// Mitsubishi GX Works2 project: ZhaoQing_OCV__Debug   PLC: Q10UDEH (continued)

Conveyor12109(ConveyorMotor:=ConveyorIO12109);
ConveyorIO12109.xForward:=M53;
ConveyorIO12109.xCWPresent:=X29;
Y22A:=ConveyorIO12109.xMotorCW;
M326:=NOT ConveyorIO12109.xEmpty;
M327:=ConveyorIO12109.xError;
ConveyorIO12109.iDeviceID:=12109;

Switch12310(ConveyorEntryIO:=ConveyorIO12110 ,
                                                        ConveyorExitIO:=ConveyorIO12117 ,
                                                        SwitchIO:=SwitchIO12310 );
SwitchIO12310.xLiftCylinderExtendButton:=M54;
SwitchIO12310.xLiftCylinderRetractButton:=M55;
Y22E:=SwitchIO12310.xLiftCylinderExtend;
Y22D:=SwitchIO12310.xLiftCylinderRetract;
SwitchIO12310.xLiftCylinderExtendDetect:=X2D;
SwitchIO12310.xLiftCylinderRetractDetect:=X2E;
ConveyorIO12110.xForward:=M56;
ConveyorIO12110.xCWPresent:=X2F OR X30;
Y22C:=ConveyorIO12110.xMotorCW;
M328:=NOT ConveyorIO12110.xEmpty;
M329:=ConveyorIO12110.xError;
ConveyorIO12110.iDeviceID:=12110;
ConveyorIO12110.tLoadDelay:=T#3s;
ConveyorIO12117.xForward:=M57;
ConveyorIO12117.xCWPresent:=X2F OR X30;
Y22F:=ConveyorIO12117.xMotorCW;
M330:=NOT ConveyorIO12117.xEmpty;
M331:=ConveyorIO12117.xError;
ConveyorIO12117.iDeviceID:=12117;

Conveyor12118(ConveyorMotor:=ConveyorIO12118);
ConveyorIO12118.xForward:=M58;
ConveyorIO12118.xCWPresent:=X31;
Y230:=conveyorIO12118.xMotorCW;
M332:=NOT ConveyorIO12118.xEmpty;
M333:=ConveyorIO12118.xError;
ConveyorIO12118.iDeviceID:=12118;

Conveyor12119(ConveyorMotor:=ConveyorIO12119);
ConveyorIO12119.xForward:=M59;
ConveyorIO12119.xCWPresent:=X32;
Y231:=conveyorIO12119.xMotorCW;
M334:=NOT ConveyorIO12119.xEmpty;
M335:=ConveyorIO12119.xError;
ConveyorIO12119.iDeviceID:=12119;
(*常温库出库分流顶升移载*)
Switch12203(ConveyorEntryIO:=ConveyorIO12142 ,
                                                        ConveyorExitIO:=ConveyorIO12203 ,
                                                        SwitchIO:=SwitchIO12203);
SwitchIO12203.xLiftCylinderExtendButton:=M60;
SwitchIO12203.xLiftCylinderRetractButton:=M61;
SwitchIO12203.xExitBarCylinderRetractButton:=M64;
Y26B:=SwitchIO12203.xExitBarCylinderRetract;
Y269:=SwitchIO12203.xLiftCylinderExtend;
Y268:=SwitchIO12203.xLiftCylinderRetract;
SwitchIO12203.xLiftCylinderExtendDetect:=X88;
SwitchIO12203.xLiftCylinderRetractDetect:=X89;
ConveyorIO12142.xForward:=M62;
ConveyorIO12142.xCWPresent:=X87;
Y281:=ConveyorIO12142.xMotorCW;
ConveyorIO12142.tLoadDelay:=T#3s;
M336:=NOT ConveyorIO12142.xEmpty;
M337:=ConveyorIO12142.xError;
ConveyorIO12142.iDeviceID:=12142;
ConveyorIO12203.xForward:=M63;
ConveyorIO12203.xCWPresent:=X87;
Y26A:=ConveyorIO12203.xMotorCW;
SwitchIO12203.xLiftCylinderExtendInit:=0;
M352:=NOT ConveyorIO12203.xEmpty;
M353:=ConveyorIO12203.xError;
ConveyorIO12203.iDeviceID:=12203;
(*常温库空框换内衬*)
Bar12326(BarCylinderIO:=BarIO12326);
BarIO12326.tLoadDelay:=T#2s;
BarIO12326.xBarCylinderButton:=M64;
BarIO12326.xPresentSwitch:=X94;
BarIO12326.xTransportMotorCWButton:=M65;
Y26E:= BarIO12326.xTransportMotorCW OR M174;
Y26C:=BarIO12326.xBarCylinder;

Switch12204(ConveyorEntryIO:=ConveyorIO12145 ,
                                                        ConveyorExitIO:=ConveyorIO12204 ,
                                                        SwitchIO:=SwitchIO12204);
SwitchIO12204.xLiftCylinderExtendButton:=M127;
SwitchIO12204.xLiftCylinderRetractButton:=M128;
Y270:=SwitchIO12204.xLiftCylinderExtend;
Y26F:=SwitchIO12204.xLiftCylinderRetract;
SwitchIO12204.xLiftCylinderExtendDetect:=X95;
SwitchIO12204.xLiftCylinderRetractDetect:=X96;
ConveyorIO12145.xForward:=M129;
ConveyorIO12145.xCWPresent:=X93;
(*Y26E:=ConveyorIO12145.xMotorCW;*)
ConveyorIO12145.tLoadDelay:=T#3s;
ConveyorIO12145.iDeviceID:=12204;
ConveyorIO12204.xForward:=M130;
ConveyorIO12204.xCWPresent:=X97;
Y271:=ConveyorIO12204.xMotorCW;
SwitchIO12204.xLiftCylinderExtendInit:=0;
M354:=NOT ConveyorIO12204.xEmpty;
M355:=ConveyorIO12204.xError;
ConveyorIO12204.iDeviceID:=12204;

Conveyor12151(ConveyorMotor:=ConveyorIO12151);
ConveyorIO12151.xForward:=M131;
ConveyorIO12151.xCWPresent:=X98;
Y272:=conveyorIO12151.xMotorCW;
M356:=NOT ConveyorIO12151.xEmpty;
M357:=ConveyorIO12151.xError;
ConveyorIO12151.iDeviceID:=12151;

Conveyor12150(ConveyorMotor:=ConveyorIO12150);
ConveyorIO12150.xForward:=M132;
ConveyorIO12150.xCWPresent:=X99;
Y273:=conveyorIO12150.xMotorCW;
M358:=NOT ConveyorIO12150.xEmpty;
M359:=ConveyorIO12150.xError;
ConveyorIO12150.iDeviceID:=12150;

Switch12328(ConveyorEntryIO:=ConveyorIO12149 ,
                                                        ConveyorExitIO:=ConveyorIO12148 ,
                                                        SwitchIO:=SwitchIO12328);
SwitchIO12328.xLiftCylinderExtendButton:=M133;
SwitchIO12328.xLiftCylinderRetractButton:=M134;
Y275:=SwitchIO12328.xLiftCylinderExtend;
Y274:=SwitchIO12328.xLiftCylinderRetract;
SwitchIO12328.xLiftCylinderExtendDetect:=X9B;
SwitchIO12328.xLiftCylinderRetractDetect:=X9C;
ConveyorIO12149.xForward:=M135;
ConveyorIO12149.xCWPresent:=X9A;
Y276:=ConveyorIO12149.xMotorCW;
ConveyorIO12149.tLoadDelay:=T#3s;
ConveyorIO12149.iDeviceID:=12148;
ConveyorIO12148.xForward:=M136;
ConveyorIO12148.xCWPresent:=X9A;
Y277:=ConveyorIO12148.xMotorCW;
M360:=NOT ConveyorIO12148.xEmpty;
M361:=ConveyorIO12148.xError;
ConveyorIO12148.iDeviceID:=12148;
SwitchIO12328.xLiftCylinderExtendInit:=0;

(*常温库去OCV线体*)
Conveyor12143(ConveyorMotor:=ConveyorIO12143);
ConveyorIO12143.xForward:=M66;
ConveyorIO12143.xCWPresent:=XA2;
Y282:=ConveyorIO12143.xMotorCW;
M338:=NOT ConveyorIO12143.xEmpty;
M339:=ConveyorIO12143.xError;
ConveyorIO12143.iDeviceID:=12143;
(*常温库OCV1顶升移载*)
Switch12330(ConveyorEntryIO:=ConveyorIO12144 ,
                                                        ConveyorExitIO:=Switch12330ConveyorOut ,
                                                        SwitchIO:=SwitchIO12330);
SwitchIO12330.xLiftCylinderExtendButton:=M67;
SwitchIO12330.xLiftCylinderRetractButton:=M68;
SwitchIO12330.xExitBarCylinderRetractButton:=M69;
Y286:=SwitchIO12330.xExitBarCylinderRetract;
Y284:=SwitchIO12330.xLiftCylinderExtend;
Y285:=SwitchIO12330.xLiftCylinderRetract;
SwitchIO12330.xLiftCylinderExtendDetect:=XA3;
SwitchIO12330.xLiftCylinderRetractDetect:=XA4;
ConveyorIO12144.xForward:=M70;
ConveyorIO12144.xCWPresent:=XA7;
Y280:=ConveyorIO12144.xMotorCW;
M340:=NOT ConveyorIO12144.xEmpty;
M341:=ConveyorIO12144.xError OR Switch12330ConveyorOut.xError;
ConveyorIO12144.iDeviceID:=12144;
ConveyorIO12144.tLoadDelay:=T#2s;
Switch12330ConveyorOut.xForward:=M178;
Switch12330ConveyorOut .xCWPresent:=XA7;
Y27C:=Switch12330ConveyorOut.xMotorCW;
Switch12330ConveyorOut.iDeviceID:=12144;

(*OCV1工位*)
Conveyor12160(ConveyorMotor:= ConveyorIO12160 );
 ConveyorIO12160.xForward:=M179;
 ConveyorIO12160.xCWPresent:=XA1;
 Y27D:= ConveyorIO12160.xMotorCW;
 M416:=NOT ConveyorIO12160.xEmpty;
 M417:=ConveyorIO12160.xError;
 ConveyorIO12160.iDeviceID:=12160;
 
(*分拣工位*)
Conveyor12146(ConveyorMotor:=ConveyorIO12146  );
ConveyorIO12146.xForward:=M71;
ConveyorIO12146.xCWPresent:=XA6;
Y283:=ConveyorIO12146.xMotorCW;
M350:=NOT ConveyorIO12146.xEmpty;
M351:=ConveyorIO12146.xError;
ConveyorIO12146.iDeviceID:=12146;

Conveyor12147(ConveyorMotor:=ConveyorIO12147);
ConveyorIO12147.xForward:=M106;
ConveyorIO12147.xCWPresent:=XA0;
Y279:=ConveyorIO12147.xMotorCW;
M342:=NOT ConveyorIO12147.xEmpty;
M343:=ConveyorIO12147.xError;
ConveyorIO12147.iDeviceID:=12147;
(*OCV2顶升移载*)
Switch12333(ConveyorEntryIO:=ConveyorIO12333 ,
                                                        ConveyorExitIO:=ConveyorIO12152 ,
                                                        SwitchIO:=SwitchIO12333);
SwitchIO12333.xLiftCylinderExtendButton:=M72;
SwitchIO12333.xLiftCylinderRetractButton:=M73;
SwitchIO12333.xEntryBarCylinderRetractButton:=M74;
Y287:=SwitchIO12333.xEntryBarCylinderRetract;
Y289:=SwitchIO12333.xLiftCylinderExtend;
Y28A:=SwitchIO12333.xLiftCylinderRetract;
SwitchIO12333.xLiftCylinderExtendDetect:=XAC;
SwitchIO12333.xLiftCylinderRetractDetect:=XAD;
ConveyorIO12333.xForward:=M75;
ConveyorIO12333.xCWPresent:=XAB;
Y288:=ConveyorIO12333.xMotorCW;
ConveyorIO12333.tLoadDelay:=T#2s;
M344:=NOT ConveyorIO12333.xEmpty;
M345:=ConveyorIO12333.xError;
ConveyorIO12333.iDeviceID:=12333;
ConveyorIO12152.xForward:=M76;
ConveyorIO12152.xCWPresent:=XAB;
(*Y28B:=ConveyorIO12152.xMotorCW;*)
Y28B:=X0FE;(*临时人工操作按钮*)
M346:=NOT ConveyorIO12152.xEmpty;
M347:=ConveyorIO12152.xError;
ConveyorIO12152.iDeviceID:=12152;

Rotor12501(ShuttleCarInOut:=RotorIO12501);
ShuttleCarCurrentPosition(XD5 OR XD6  ,XD5 ,XD6, FALSE, RotorIO12501.iCurrentPos);
RotorIO12501.xReady:=XB9;
RotorIO12501.xForward:=M158;
RotorIO12501.xBackward:=M159;
RotorIO12501.xPosLimit:=XD7;
RotorIO12501.xNegLimit:=XD8;
Y2A9:=RotorIO12501.xCW;
Y2AA:=RotorIO12501.xCCW;
Y2AE:=RotorIO12501.xBrake;

Conveyor12501(ConveyorMotor:=ConveyorIO12501);
ConveyorIO12501.xForward:=M160;
ConveyorIO12501.xBackward:=M161;
ConveyorIO12501.xCWPresent:=XD9;
ConveyorIO12501.xCCWPresent:=XDA;
Y2AF:=ConveyorIO12501.xMotorCW;
Y2B0:=ConveyorIO12501.xMotorCCW;
M348:=NOT ConveyorIO12501.xEmpty;
M349:=ConveyorIO12501.xError;
ConveyorIO12501.iDeviceID:=12501;

Conveyor12154(ConveyorMotor:=ConveyorIO12154);
ConveyorIO12154.xForward:=M168;
ConveyorIO12154.xCWPresent:=XB8;
Y28F:=ConveyorIO12154.xMotorCW;
M383:=NOT ConveyorIO12154.xEmpty;
M384:=ConveyorIO12154.xError;
ConveyorIO12154.iDeviceID:=12154;

(******OCV入库线体******)

(*常温库入库前端线体*)
Conveyor12159(ConveyorMotor:=ConveyorIO12159);
ConveyorIO12159.xForward:=M119;
ConveyorIO12159.xCWPresent:=XE1;
Y2B8:=ConveyorIO12159.xMotorCW;
M365:=NOT ConveyorIO12159.xEmpty;
M366:=ConveyorIO12159.xError;
ConveyorIO12159.iDeviceID:=12159;

(*常温库入库前顶升移载*)
Switch12337(ConveyorEntryIO:= ConveyorIO12158 ,ConveyorExitIO:= ConveyorIO12157 ,SwitchIO:= SwitchIO12337 );
SwitchIO12337.xLiftCylinderExtendButton:=M120;
SwitchIO12337.xLiftCylinderRetractButton:=M121;
Y2B6:=SwitchIO12337.xLiftCylinderExtend;
Y2B5:=SwitchIO12337.xLiftCylinderRetract;
SwitchIO12337.xLiftCylinderExtendDetect:=XDE;
SwitchIO12337.xLiftCylinderRetractDetect:=XDF;
ConveyorIO12158.xForward:=M122;
ConveyorIO12158.xCWPresent:=XDD;
Y2B7:=ConveyorIO12158.xMotorCW;
ConveyorIO12158.tLoadDelay:=T#2s;
M367:=NOT ConveyorIO12158.xEmpty;
M368:=ConveyorIO12158.xError;
ConveyorIO12158.iDeviceID:=12158;
ConveyorIO12157.xForward:=M123;
ConveyorIO12157.xCWPresent:=XDD;
Y2B4:=ConveyorIO12157.xMotorCW;
M369:=NOT ConveyorIO12157.xEmpty;
M370:=ConveyorIO12157.xError;
ConveyorIO12157.iDeviceID:=12157;

Conveyor12156(ConveyorMotor:=ConveyorIO12156);
ConveyorIO12156.xForward:=M116;
ConveyorIO12156.xCWPresent:=XDC;
Y2B2:=ConveyorIO12156.xMotorCW;
M371:=NOT ConveyorIO12156.xEmpty;
M372:=ConveyorIO12156.xError;
ConveyorIO12156.iDeviceID:=12156;

Conveyor12155(ConveyorMotor:=ConveyorIO12155);
ConveyorIO12155.xForward:=M117;
ConveyorIO12155.xCWPresent:=XDB;
Y2B3:=ConveyorIO12155.xMotorCW;
M373:=NOT ConveyorIO12155.xEmpty;
M374:=ConveyorIO12155.xError;
ConveyorIO12155.iDeviceID:=12155;

Conveyor12141(ConveyorMotor:=ConveyorIO12141);
ConveyorIO12141.xForward:=M124;
ConveyorIO12141.xCWPresent:=XF0;
Y2C5:=ConveyorIO12141.xMotorCW;
M375:=NOT ConveyorIO12141.xEmpty;
M376:=ConveyorIO12141.xError;
ConveyorIO12141.iDeviceID:=12141;
(******常温库1巷道入库******)
Switch12321(ConveyorEntryIO:=ConveyorIO12321 ,
                                                        ConveyorExitIO:=ConveyorIO12140 ,
                                                        SwitchIO:=SwitchIO12321);
SwitchIO12321.xLiftCylinderExtendButton:=M77;
SwitchIO12321.xLiftCylinderRetractButton:=M78;
SwitchIO12321.xExitBarCylinderRetractButton:=M79;
Y267:=SwitchIO12321.xExitBarCylinderRetract OR m_iSwitch12321Select=2 OR M173;
Y266:=SwitchIO12321.xExitBarCylinderRetract OR M173;
Y265:=SwitchIO12321.xLiftCylinderExtend;
Y264:=SwitchIO12321.xLiftCylinderRetract;
SwitchIO12321.xLiftCylinderExtendDetect:=X7C;
SwitchIO12321.xLiftCylinderRetractDetect:=X7D;
ConveyorIO12321.xForward:=M80;
ConveyorIO12321.xCWPresent:=((m_iSwitch12321Select=1 OR m_iSwitch12321Select=0) AND   X7E) OR (m_iSwitch12321Select=2 AND X79);
Y263:=ConveyorIO12321.xMotorCW;
ConveyorIO12321.tLoadDelay:=T#3s;
ConveyorIO12321.iDeviceID:=12321;
ConveyorIO12140.xForward:=M81;
ConveyorIO12140.xCWPresent:=((m_iSwitch12321Select=1 OR m_iSwitch12321Select=0) AND   X7E) OR (m_iSwitch12321Select=2 AND X79);
Y261:=ConveyorIO12140.xMotorCW;
M377:=NOT ConveyorIO12140.xEmpty;
M378:=ConveyorIO12140.xError;
ConveyorIO12140.iDeviceID:=12140;

Conveyor12138(ConveyorMotor:=ConveyorIO12138);
ConveyorIO12138.xForward:=M82;
ConveyorIO12138.xCWPresent:=X71;
Y25F:=ConveyorIO12138.xMotorCW;
ConveyorIO12138.tLoadDelay:=t#2s;
M379:=NOT ConveyorIO12138.xEmpty;
M380:=ConveyorIO12138.xError;
ConveyorIO12138.iDeviceID:=12138;

Conveyor12139(ConveyorMotor:=ConveyorIO12139);
ConveyorIO12139.xForward:=M83;
ConveyorIO12139.xCWPresent:=X73;
Y260:=ConveyorIO12139.xMotorCW;
ConveyorIO12139.tLoadDelay:=t#2s;
M381:=NOT ConveyorIO12139.xEmpty;
M382:=ConveyorIO12139.xError;
ConveyorIO12139.iDeviceID:=12139;

Cylinder12320(ShuttleCarInOut:= CylinderIO12320 );
ShuttleCarCurrentPosition( X75 OR X76 ,X76 ,X75, FALSE, CylinderIO12320.iCurrentPos );
CylinderIO12320.xForward:=M102;
CylinderIO12320.xBackward:=M103;
Y25E:=CylinderIO12320.xCW;
Y25D:=CylinderIO12320.xCCW;
CylinderIO12320.xCylinder:=1;
CylinderIO12320.xPresentDetect1:=X74;
CylinderIO12320.xPresentDetect2:=X72;

(******常温库2巷道入库******)
Conveyor12137(ConveyorMotor:=ConveyorIO12137);
ConveyorIO12137.xForward:=M84;
ConveyorIO12137.xCWPresent:=X70;
Y25C:=ConveyorIO12137.xMotorCW;
ConveyorIO12137.iDeviceID:=12137;
M385:=NOT ConveyorIO12137.xEmpty;
M386:=ConveyorIO12137.xError;
ConveyorIO12137.iDeviceID:=12137;

Conveyor12136(ConveyorMotor:=ConveyorIO12136);
ConveyorIO12136.xForward:=M85;
ConveyorIO12136.xCWPresent:=X6F;
Y25B:=ConveyorIO12136.xMotorCW;
M387:=NOT ConveyorIO12136.xEmpty;
M388:=ConveyorIO12136.xError;
ConveyorIO12136.iDeviceID:=12136;


Switch12317(ConveyorEntryIO:=ConveyorIO12135 ,
                                                        ConveyorExitIO:=ConveyorIO12134 ,
                                                        SwitchIO:=SwitchIO12317);
SwitchIO12317.xLiftCylinderExtendButton:=M86;
SwitchIO12317.xLiftCylinderRetractButton:=M87;
SwitchIO12317.xExitBarCylinderRetractButton:=M88;
Y259:=SwitchIO12317.xExitBarCylinderRetract OR m_iSwitch12317Select=2 ;
Y256:=SwitchIO12317.xExitBarCylinderRetract ;
Y258:=SwitchIO12317.xLiftCylinderExtend;
Y257:=SwitchIO12317.xLiftCylinderRetract;
SwitchIO12317.xLiftCylinderExtendDetect:=X6A;
SwitchIO12317.xLiftCylinderRetractDetect:=X6B;
ConveyorIO12135.xForward:=M89;
ConveyorIO12135.xCWPresent:=((m_iSwitch12317Select=1 OR m_iSwitch12317Select=0) AND   X6E) OR (m_iSwitch12317Select=2 AND X67);
Y25A:=ConveyorIO12135.xMotorCW;
ConveyorIO12135.tLoadDelay:=T#3s;
M389:=NOT ConveyorIO12135.xEmpty;
M390:=ConveyorIO12135.xError;
ConveyorIO12135.iDeviceID:=12135;
ConveyorIO12134.xForward:=M90;
ConveyorIO12134.xCWPresent:=((m_iSwitch12317Select=1 OR m_iSwitch12317Select=0) AND   X6E) OR (m_iSwitch12317Select=2 AND X67);
Y255:=ConveyorIO12134.xMotorCW;
M391:=NOT ConveyorIO12134.xEmpty;
M392:=ConveyorIO12134.xError;
ConveyorIO12134.iDeviceID:=12134;

Conveyor12132(ConveyorMotor:=ConveyorIO12132);
ConveyorIO12132.xForward:=M91;
ConveyorIO12132.xCWPresent:=X5F;
Y253:=ConveyorIO12132.xMotorCW;
ConveyorIO12132.tLoadDelay:=t#2s;
M393:=NOT ConveyorIO12132.xEmpty;
M394:=ConveyorIO12132.xError;
ConveyorIO12132.iDeviceID:=12132;

Conveyor12133(ConveyorMotor:=ConveyorIO12133);
ConveyorIO12133.xForward:=M92;
ConveyorIO12133.xCWPresent:=X61;
Y254:=ConveyorIO12133.xMotorCW;
ConveyorIO12133.tLoadDelay:=t#2s;
M395:=NOT ConveyorIO12133.xEmpty;
M396:=ConveyorIO12133.xError;
ConveyorIO12133.iDeviceID:=12133;

Cylinder12316(ShuttleCarInOut:= CylinderIO12316 );
ShuttleCarCurrentPosition( X63 OR X64 ,X64 ,X63, FALSE, CylinderIO12316 .iCurrentPos );
CylinderIO12316 .xForward:=M125;
CylinderIO12316 .xBackward:=M126;
Y252:=CylinderIO12316 .xCW;
Y251:=CylinderIO12316 .xCCW;
CylinderIO12316.xCylinder:=1;
CylinderIO12316.xPresentDetect1:=X62;
CylinderIO12316.xPresentDetect2:=X60;
(******常温库3巷道入库******)
Conveyor12131(ConveyorMotor:=ConveyorIO12131);
ConveyorIO12131.xForward:=M93;
ConveyorIO12131.xCWPresent:=X5E;
Y24E:=ConveyorIO12131.xMotorCW;
M397:=NOT ConveyorIO12131.xEmpty;
M398:=ConveyorIO12131.xError;
ConveyorIO12131.iDeviceID:=12131;

Conveyor12130(ConveyorMotor:=ConveyorIO12130);
ConveyorIO12130.xForward:=M94;
ConveyorIO12130.xCWPresent:=X5D;
Y24F:=ConveyorIO12130.xMotorCW;
M399:=NOT ConveyorIO12130.xEmpty;
M400:=ConveyorIO12130.xError;
ConveyorIO12130.iDeviceID:=12130;

Switch12314(ConveyorEntryIO:=ConveyorIO12129 ,
                                                        ConveyorExitIO:=ConveyorIO12128 ,
                                                        SwitchIO:=SwitchIO12314);
SwitchIO12314.xLiftCylinderExtendButton:=M95;
SwitchIO12314.xLiftCylinderRetractButton:=M96;
SwitchIO12314.xExitBarCylinderRetractButton:=M97;
Y24D:=SwitchIO12314.xExitBarCylinderRetract OR m_iSwitch12314Select=2 ;
Y24C:=SwitchIO12314.xLiftCylinderExtend;
Y24B:=SwitchIO12314.xLiftCylinderRetract;
SwitchIO12314.xLiftCylinderExtendDetect:=X58;
SwitchIO12314.xLiftCylinderRetractDetect:=X59;
ConveyorIO12129.xForward:=M98;
ConveyorIO12129.xCWPresent:=((m_iSwitch12314Select=1 OR m_iSwitch12314Select=0) AND   X5C) OR (m_iSwitch12314Select=2 AND X57);
Y250:=ConveyorIO12129.xMotorCW;
ConveyorIO12129.tLoadDelay:=T#3s;
M401:=NOT ConveyorIO12129.xEmpty;
M402:=ConveyorIO12129.xError;
ConveyorIO12129.iDeviceID:=12129;
ConveyorIO12128.xForward:=M99;
ConveyorIO12128.xCWPresent:=((m_iSwitch12314Select=1 OR m_iSwitch12314Select=0) AND   X5C) OR (m_iSwitch12314Select=2 AND X57);
Y24A:=ConveyorIO12128.xMotorCW;
ConveyorIO12128.iDeviceID:=12128;
M403:=NOT ConveyorIO12128.xEmpty;
M404:=ConveyorIO12128.xError;

Conveyor12126(ConveyorMotor:=ConveyorIO12126);
ConveyorIO12126.xForward:=M100;
ConveyorIO12126.xCWPresent:=X4F;
ConveyorIO12126.tLoadDelay:=t#2s;
Y248:=ConveyorIO12126.xMotorCW;
M405:=NOT ConveyorIO12126.xEmpty;
M406:=ConveyorIO12126.xError;
ConveyorIO12126.iDeviceID:=12126;

Conveyor12127(ConveyorMotor:=ConveyorIO12127);
ConveyorIO12127.xForward:=M101;
ConveyorIO12127.xCWPresent:=X51;
Y249:=ConveyorIO12127.xMotorCW;
ConveyorIO12127.tLoadDelay:=t#2s;
M407:=NOT ConveyorIO12127.xEmpty;
M408:=ConveyorIO12127.xError;
ConveyorIO12127.iDeviceID:=12127;

Cylinder12313(ShuttleCarInOut:= CylinderIO12313 );
ShuttleCarCurrentPosition( X53 OR X54 ,X54 ,X53, FALSE, CylinderIO12313 .iCurrentPos );
CylinderIO12313 .xForward:=M104;
CylinderIO12313 .xBackward:=M105;
Y247:=CylinderIO12313 .xCW;
Y246:=CylinderIO12313 .xCCW;
CylinderIO12313.xCylinder:=1;
CylinderIO12313.xPresentDetect1:=X52;
CylinderIO12313.xPresentDetect2:=X50;

(**************************)
IF g_xManual THEN
	D3165:=0;
	D3185:=0;
	D3160:=0;
	D3161:=0;
	D3162:=0;
	D3180:=0;
	D3181:=0;
	D3182:=0;
	D3200:=0;
	D3201:=0;
	D3202:=0;		
	D3330:=0;
	D3325:=0;
END_IF;
IF g_xAuto THEN
(*	"OCV前分流
4007"	2330	5	分流方向	2330	"0：复位
1：读码失败
2：流向OCV1，
3：流向OCV2"	3330	5	有板状态	3330	1：无板，2：有板*)
IF ConveyorIO12125.xEmpty=0 THEN
	D3330:=2;
ELSE
	D3330:=1;	
END_IF;
IF ldp(TRUE,  D2330>1) THEN
	ConveyorIO12125.iProductCategory:=D2330;
END_IF;
(*"常温入库前分流（OCV1后）
4006"	2325	5	分流方向	2325	"0：复位
1：读码失败
2：流向C1库，
3：流向C2库
4：流向C3库"	3325	5	有板状态	3325	1：无板，2：有板*)
IF ConveyorIO12155.xEmpty=0 THEN
	D3325:=2;
ELSE
	D3325:=1;
END_IF;
IF LDP(TRUE,D2325>1) THEN
	ConveyorIO12155.iProductCategory:=D2325;
END_IF;
(*	"C1库入口(OCV1后）
2013
（出入口编号3）"	2160	5				3160	5	位置1有板状态	3160	1：无板，2：有板
								位置2有板状态	3161	1：无板，2：有板
								手动入库请求	3162	1:复位，2：请求入库*)
	IF CylinderIO12320.iCurrentPos=2 AND CylinderIO12320.xPresentDetect1 AND NOT M170 THEN
		D3160:=2;
	ELSIF M170 THEN
		D3160:=0;
	ELSE
		D3160:=1;
	END_IF;
	IF CylinderIO12320.iCurrentPos=2 AND CylinderIO12320.xPresentDetect2 AND NOT M170 THEN
		D3161:=2;
	ELSIF M170 THEN
		D3161:=0;
	ELSE
		D3161:=1;
	END_IF;	
    IF  g_xImport1Force AND (CylinderIO12320.xPresentDetect2 OR CylinderIO12320.xPresentDetect1)THEN
  		D3162:=2;
  	END_IF;	
	IF D2160 =2 THEN  (*Reset request*)
		D3162:=1;
    END_IF;	  
(*"C2库入口(OCV1后）
2017
（出入口编号3）"	2180	5				3180	5	位置1有板状态	3180	1：无板，2：有板
								位置2有板状态	3181	1：无板，2：有板
								手动入库请求	3182	1:复位，2：请求入库*)
	IF CylinderIO12316.iCurrentPos=2 AND CylinderIO12316.xPresentDetect1 AND NOT M171 THEN
		D3180:=2;
	ELSIF M171 THEN
		D3180:=0;
		ELSE
		D3180:=1;
	END_IF;
	IF CylinderIO12316.iCurrentPos=2 AND CylinderIO12316.xPresentDetect2 AND NOT  M171 THEN
		D3181:=2;
	ELSIF M171 THEN
		D3181:=0;		
	ELSE
		D3181:=1;
	END_IF;	
    IF  g_xImport2Force AND (CylinderIo12316.xPresentDetect1	OR CylinderIO12316.xPresentDetect2) THEN
  		D3182:=2;
  	END_IF;
	IF D2180=2 THEN
		D3182:=1;
    END_IF;	
(*	"C3库入口(OCV1后）
2021
（出入口编号3）"	2200	5				3200	5	位置1有板状态	3200	1：无板，2：有板
								位置2有板状态	3201	1：无板，2：有板
								手动入库请求	3202	1:复位，2：请求入库*)
	IF CylinderIO12313.iCurrentPos=2 AND CylinderIO12313.xPresentDetect1 AND NOT M172 THEN
		D3200:=2;
	ELSIF M172 THEN
		D3200:=0;
	ELSE
		D3200:=1;
	END_IF;
	IF CylinderIO12313.iCurrentPos=2 AND CylinderIO12313.xPresentDetect2 AND NOT M172 THEN
		D3201:=2;
	ELSIF M172 THEN
		D3201:=0;
	ELSE
		D3201:=1;
	END_IF;	
    IF  g_xImport3Force AND (CylinderIO12313.xPresentDetect1 OR CylinderIO12313.xPresentDetect2) THEN
  		D3202:=2;
  	END_IF;
	IF D2200=2 THEN
		D3202:=1;
    END_IF;	

	(*与上位机接口程序
	"C1库出口(产品出库)
2014
出库完成状态	2165	"1：复位2：出库完成
出口状态	3165	"1:禁止出库2:允许出库"
1线堆积状态	3166	"1：正常2:堆积 "
2线堆积状态	3167	"1：正常2:堆积 "
3线堆积状态	3168	"1：正常2:堆积 "
    (**************************)
    IF NOT X41 AND NOT X42 AND CylinderIO12309.iCurrentPos=2 AND NOT M175 THEN
    	D3165:=2;
    ELSIF M175 THEN
    	D3165:=0;
    ELSE
    	D3165:=1;
    END_IF;
   IF D2165=2 THEN
   		m_xTS1ExportPermit:=1;
   ELSE
   		m_xTS1ExportPermit:=0;
   END_IF;
(*"C2库出口(产品出库)
2018
（出入口编号4）"	2185	5	出库完成状态	2185	"1：复位
2：出库完成 "	3185	5	出口状态	3185	"1:禁止出库
2:允许出库"
								1线堆积状态	3186	"1：正常
2:堆积 "
								2线堆积状态	3187	"1：正常
2:堆积 "
								3线堆积状态	3188	"1：正常
2:堆积 "
*)
    IF NOT X33 AND NOT X34 AND CylinderIO12308.iCurrentPos=2 AND NOT M176 THEN
    	D3185:=2;
    ELSIF M176 THEN
    	D3185:=0;
    ELSE
    	D3185:=1;
    END_IF;
   IF D2185=2 THEN
   		m_xTS2ExportPermit:=1;
   ELSE
   		m_xTS2ExportPermit:=0;
   END_IF;
   (**************************)
 (*  "C3库出口(产品出口)
2022
（出入口编号4）"	2205	5	出库完成状态	2205	"1：复位
2：出库完成 "	3205	5	出口状态	3205	"1:禁止出库
2:允许出库"
								1线堆积状态	3206	"1：正常
2:堆积 "
								2线堆积状态	3207	"1：正常
2:堆积 "
								3线堆积状态	3208	"1：正常
2:堆积 "*)
   IF NOT CylinderIO12307.xPresentDetect1 
   	AND NOT CylinderIO12307.xPresentDetect2 
   	AND CylinderIO12307.iCurrentPos=2
   	AND NOT M177  THEN
      	D3205:=2;
   ELSIF M177  THEN
   	D3205:=0;
   	ELSE
    	D3205:=1;
    END_IF; 	
   IF D2205=2 THEN
   		m_xTS3ExportPermit:=1;
   ELSE
   		m_xTS3ExportPermit:=0;
   END_IF;


    (**************常温库3巷道出库************) 
	IF NOT CylinderIO12307.xPresentDetect1 
		AND NOT CylinderIO12307.xPresentDetect2
		AND ConveyorIO12108.xEmpty 
		AND ConveyorIO12109.xEmpty 
		AND NOT ConveyorIO12108.xBusy 
		AND NOT ConveyorIO12109.xBusy THEN
		CylinderIO12307.xMDIExe:=1;
		CylinderIO12307.iDestinationPos:=2;
	END_IF;
	IF (m_xTS3ExportPermit=1 OR M164) AND ( CylinderIO12307.xPresentDetect1  OR CylinderIO12307.xPresentDetect2) THEN
		CylinderIO12307.xMDIExe:=1;
		CylinderIO12307.iDestinationPos:=1;
	END_IF;
	
	IF CylinderIO12307.iCurrentPos=1 AND CylinderIO12307.xPresentDetect1 THEN
		ConveyorIO12108.xLoad:=1;
	ELSE
		ConveyorIO12108.xLoad:=0;
	END_IF;
	IF CylinderIO12307.iCurrentPos=1 AND CylinderIO12307.xPresentDetect2 THEN
		ConveyorIO12109.xLoad:=1;
	ELSE
		ConveyorIO12109.xLoad:=0;	
	END_IF;	
	SwitchIO12310.xEntryEnable:=(ConveyorIO12108.xNextRun OR ConveyorIO12109.xNextRun) AND ConveyorIO12117.xEmpty ;
    ConveyorIO12108.xUnload:=ConveyorIO12110.xEmpty ;
    SwitchIO12310.xSwithEnable:=1;
     SwitchIO12310.xLiftCylinderExtendInit:=1;
    SwitchIO12310.xExitEnable:=ConveyorIo12118.xEmpty;
    IF ConveyorIO12108.xEmpty AND conveyorIO12117.xEmpty AND NOT ConveyorIO12108.xBusy THEN
    	ConveyorIO12109.xUnload:=ConveyorIO12110.xEmpty AND ConveyorIO12117.xEmpty ;
    ELSE
    	ConveyorIO12109.xUnload:=0;
    END_IF;
    ConveyorIO12118.xLoad:=ConveyorIO12117 .xNextRun;
    ConveyorIO12118.xUnload:=ConveyorIO12119.xEmpty;
    ConveyorIO12119.xLoad:=ConveyorIO12118.xNextRun;
    (*汇流点防止碰撞*)
    ConveyorIO12119.xUnload:=ConveyorIO12120.xEmpty AND m_xSwitch12311Task=3;   
     IF m_xSwitch12311Task=3 OR  m_xSwitch12311Task=0 THEN
    	SwitchIO12311.xLiftCylinderExtendInit:=0;
    END_IF;
    ConveyorIO12120.xLoad:=ConveyorIO12119.xNextRun;    
    
    (**************常温库2巷道出库************) 
	IF NOT X33 
		AND NOT X34 
		AND ConveyorIO12111.xEmpty 
		AND ConveyorIO12112.xEmpty 
		AND NOT ConveyorIO12111.xBusy 
		AND NOT ConveyorIO12112.xBusy THEN
		CylinderIO12308.xMDIExe:=1;
		CylinderIO12308.iDestinationPos:=2;
	END_IF;
	IF (m_xTS2ExportPermit=1 OR M163) AND ( X33 OR X34) THEN
		CylinderIO12308.xMDIExe:=1;
		CylinderIO12308.iDestinationPos:=1;
	END_IF;
	
	IF CylinderIO12308.iCurrentPos=1 AND X34 THEN
		ConveyorIO12111.xLoad:=1;
	ELSE
		ConveyorIO12111.xLoad:=0;
	END_IF;
	IF CylinderIO12308.iCurrentPos=1 AND X33 THEN
		ConveyorIO12112.xLoad:=1;
	ELSE
		ConveyorIO12112.xLoad:=0;	
	END_IF;	
		Switch12311Priority(xCondition1:=NOT  ConveyorIO12111.xEmpty ,
	                                       xCondition2:= NOT  ConveyorIO12112.xEmpty ,
	                                       xCondition3:= NOT  ConveyorIO12119.xEmpty,
	                                       xCondition4:= FALSE ,
	                                       xCondition5:= FALSE ,
	                                       xTaskComplete:=LDF (TRUE,ConveyorIO12120.xEmpty=0),
	                                       xReset:= g_xResetSingle AND (g_iDeviceIDSelect=12120 OR g_iDeviceIDSelect=12113),
	                                       iPriority:= m_xSwitch12311Task);
	SwitchIO12311.xEntryEnable:=(ConveyorIO12111.xNextRun AND m_xSwitch12311Task=1) OR (ConveyorIO12112.xNextRun AND m_xSwitch12311Task=2);
    ConveyorIO12111.xUnload:=ConveyorIO12113.xEmpty AND ConveyorIO12120.xEmpty AND m_xSwitch12311Task=1 ;    
    IF m_xSwitch12311Task=1 OR  m_xSwitch12311Task=2 THEN
  	  SwitchIO12311.xLiftCylinderExtendInit:=1;
  	  SwitchIO12311.xSwithEnable:=1;
    ELSE
       SwitchIO12311.xSwithEnable:=0;
    END_IF;
    SwitchIO12311.xExitEnable:=ConveyorIo12121.xEmpty;

    	ConveyorIO12112.xUnload:=ConveyorIO12113.xEmpty AND ConveyorIO12120.xEmpty AND m_xSwitch12311Task=2;
(*******************************************)
	ConveyorIO12120.xUnload:=ConveyorIO12121.xEmpty;
    ConveyorIO12121.xLoad:=ConveyorIO12120 .xNextRun;
    ConveyorIO12121.xUnload:=ConveyorIO12122.xEmpty;
    ConveyorIO12122.xLoad:=ConveyorIO12121.xNextRun;
    IF m_xSwitch12312Task=3 OR m_xSwitch12312Task=0 THEN
    	SwitchIO12312.xLiftCylinderExtendInit:=0;
    END_IF;
    (*汇流点防止碰撞*)
    ConveyorIO12122.xUnload:=ConveyorIO12123.xEmpty AND m_xSwitch12312Task=3 ; (*1巷道出库顶升移载为空*)
    ConveyorIO12123.xLoad:=ConveyorIO12122.xNextRun;
  (**************常温库1巷道出库************) 
	IF NOT X41 
		AND NOT X42 
		AND ConveyorIO12114.xEmpty 
		AND ConveyorIO12115.xEmpty 
		AND NOT ConveyorIO12114.xBusy
		AND NOT ConveyorIO12115.xBusy THEN
		CylinderIO12309.xMDIExe:=1;
		CylinderIO12309.iDestinationPos:=2;
	END_IF;
	IF (m_xTS1ExportPermit=1 OR M162) AND  (X41 OR X42) THEN (*M162强制出库*)
		CylinderIO12309.xMDIExe:=1;
		CylinderIO12309.iDestinationPos:=1;
	END_IF;
	
	IF CylinderIO12309.iCurrentPos=1 AND X41 THEN
		ConveyorIO12114.xLoad:=1;
	ELSE
		ConveyorIO12114.xLoad:=0;
	END_IF;
	IF CylinderIO12309.iCurrentPos=1  AND X42 THEN
		ConveyorIO12115.xLoad:=1;
	ELSE
		ConveyorIO12115.xLoad:=0;	
	END_IF;
	Switch12312Priority(xCondition1:=NOT  ConveyorIO12114.xEmpty ,
	                                       xCondition2:= NOT  ConveyorIO12115.xEmpty ,
	                                       xCondition3:= NOT  ConveyorIO12122.xEmpty,
	                                       xCondition4:= FALSE ,
	                                       xCondition5:= FALSE ,
	                                       xTaskComplete:=LDF (TRUE,ConveyorIO12123.xEmpty=0),
	                                       xReset:= g_xResetSingle AND (g_iDeviceIDSelect=12123 OR g_iDeviceIDSelect=12116),
	                                       iPriority:= m_xSwitch12312Task );
	SwitchIO12312.xEntryEnable:=(ConveyorIO12114.xNextRun  AND m_xSwitch12312Task=1)  OR (ConveyorIO12115.xNextRun AND m_xSwitch12312Task=2) ;
    ConveyorIO12114.xUnload:=ConveyorIO12116.xEmpty AND ConveyorIO12123.xEmpty  AND m_xSwitch12312Task=1 ;
    IF m_xSwitch12312Task=1 OR  m_xSwitch12312Task=2 THEN
  	  SwitchIO12312.xLiftCylinderExtendInit:=1;
  	  SwitchIO12312.xSwithEnable:=1;
    ELSE
      SwitchIO12312.xSwithEnable:=0;
    END_IF;
    (*SwitchIO12312.xExitEnable:=ConveyorIo12124.xEmpty;*)
    	ConveyorIO12115.xUnload:=ConveyorIO12116.xEmpty AND ConveyorIO12123.xEmpty AND m_xSwitch12312Task=2;
    (*******************************************************************)
    ConveyorIO12123.xUnload:=ConveyorIo12124.xEmpty ;
    ConveyorIO12124.xLoad:=ConveyorIO12123 .xNextRun;
    ConveyorIO12124.xUnload:=ConveyorIO12125.xEmpty;
    ConveyorIO12125.xLoad:=ConveyorIO12124.xNextRun;
     ConveyorIO12125.xUnload:=ConveyorIO12142.xEmpty AND  ConveyorIO12125.iProductCategory>1;
     (*触摸屏上计数与清零程序*)
     IF LDF(TRUE,ConveyorIO12125.xEmpty) THEN
     	D10:=D10+1;
     END_IF;
     IF M167 THEN
     	D10:=0;
     END_IF;